HMI tags "DB_SDC_ERROR_STAT"
   "SDC\DB_SDC_ERROR_STAT\_Byte_DB_SDC_ERROR_STAT.F_STAT[XX5].EMS_TS_STAT_VAL.ERROR" : Int, internal   // Fehlernummer / Error number
   "SDC\DB_SDC_ERROR_STAT\_Byte_DB_SDC_ERROR_STAT.F_STAT[XX8].F" : Int, internal   // Fehler SDC + EMS Zusammenfassung / Fault SDC + EMS Summary
   "SDC\DB_SDC_ERROR_STAT\_Byte_DB_SDC_ERROR_STAT.F_STAT[X10].EMS_TS_STAT_VAL.DRIVE_POS_PERC" : Int, internal   // Position [% of Start End Section]
   "SDC\DB_SDC_ERROR_STAT\_Byte_DB_SDC_ERROR_STAT.F_STAT[XX9].F" : Int, internal   // Fehler SDC + EMS Zusammenfassung / Fault SDC + EMS Summary
   "SDC\DB_SDC_ERROR_STAT\_Byte_DB_SDC_ERROR_STAT.F_STAT[XX6].F_DATE" : Int, internal   // Fehler Zeit / Fault Time
   "SDC\DB_SDC_ERROR_STAT\DB_SDC_ERROR_STAT.F_STAT[XX7].EMS_TS_STAT_VAL.DRIVE_POS" : DInt AT %DB0.DBD0, 1 s   // Antriebsposition in mm / Drive position in mm
   "DB_SDC_ERRORS_STAT_HEADER.FAULT_PRO_SEITE_HMI" : Int = PLC DB_SDC_ERRORS_STAT.HEADER.FAULT_PRO_SEITE_HMI AT %DB3724.DBW10, 1 s   // Reserve
   "SDC\DB_SDC_ERROR_STAT\DB_SDC_ERROR_STAT.F_STAT[XX8].EMS_TS_STAT_VAL.DRIVE_POS" : DInt AT %DB0.DBD0, 1 s   // Antriebsposition in mm / Drive position in mm
   "SDC\DB_SDC_ERROR_STAT\DB_SDC_ERROR_STAT.F_STAT[XX8].EMS_TS_STAT_VAL.SEK" : Int AT %DB0.DBW0, 1 s   // Sektion
   "SDC\DB_SDC_ERROR_STAT\_Byte_DB_SDC_ERROR_STAT.F_STAT[XX1].EMS_TS_STAT_VAL.EMS_ID" : Int, internal   // EMS ID Nummer / EMS ID Number
   "SDC\DB_SDC_ERROR_STAT\DB_SDC_ERROR_STAT.F_STAT[XX5].EMS_TS_STAT_VAL.DRIVE_POS" : DInt AT %DB0.DBD0, 1 s   // Antriebsposition in mm / Drive position in mm
   "SDC\DB_SDC_ERROR_STAT\DB_SDC_ERROR_STAT.F_STAT[XX3].F_DATE" : Date_And_Time AT %DB0.DBX0.0, 1 s   // Fehler Zeit / Fault Time
   "SDC\DB_SDC_ERROR_STAT\_Byte_DB_SDC_ERROR_STAT.F_STAT[XX9].EMS_TS_STAT_VAL.TILT_POS" : Int, internal   // Tilt angle in degrees
   "SDC\DB_SDC_ERROR_STAT\DB_SDC_ERROR_STAT.F_STAT[XX7].F_DATE" : Date_And_Time AT %DB0.DBX0.0, 1 s   // Fehler Zeit / Fault Time
   "SDC\DB_SDC_ERROR_STAT\DB_SDC_ERROR_STAT.F_STAT[XX1].F_DATE" : Date_And_Time AT %DB0.DBX0.0, 1 s   // Fehler Zeit / Fault Time
   "SDC\DB_SDC_ERROR_STAT\DB_SDC_ERROR_STAT.F_STAT[XX4].EMS_TS_STAT_VAL.DRIVE_POS_PERC" : Int AT %DB0.DBW0, 1 s   // Position [% of Start End Section]
   "SDC\DB_SDC_ERROR_STAT\_Byte_DB_SDC_ERROR_STAT.F_STAT[XX6].EMS_TS_STAT_VAL.SEK" : Int, internal   // Sektion
   "SDC\DB_SDC_ERROR_STAT\_Byte_DB_SDC_ERROR_STAT.F_STAT[XX5].EMS_TS_STAT_VAL.PROFIL" : Int, internal   // Profile
   "SDC\DB_SDC_ERROR_STAT\DB_SDC_ERROR_STAT.F_STAT[XX5].EMS_TS_STAT_VAL.SEK" : Int AT %DB0.DBW0, 1 s   // Sektion
   "SDC\DB_SDC_ERROR_STAT\DB_SDC_ERROR_STAT.F_STAT[XX6].EMS_TS_STAT_VAL.PROFIL" : Int AT %DB0.DBW0, 1 s   // Profile
   "SDC\DB_SDC_ERROR_STAT\_Byte_DB_SDC_ERROR_STAT.F_STAT[XX8].EMS_TS_STAT_VAL.EMS_ID" : Int, internal   // EMS ID Nummer / EMS ID Number
   "SDC\DB_SDC_ERROR_STAT\_Byte_DB_SDC_ERROR_STAT.F_STAT[XX6].F" : Int, internal   // Fehler SDC + EMS Zusammenfassung / Fault SDC + EMS Summary
   "SDC\DB_SDC_ERROR_STAT\_Byte_DB_SDC_ERROR_STAT.F_STAT[XX5].EMS_TS_STAT_VAL.TILT_POS" : Int, internal   // Tilt angle in degrees
   "SDC\DB_SDC_ERROR_STAT\_Byte_DB_SDC_ERROR_STAT.F_STAT[XX2].EMS_TS_STAT_VAL.SEK" : Int, internal   // Sektion
   "SDC\DB_SDC_ERROR_STAT\DB_SDC_ERROR_STAT.F_STAT[XX5].F" : Word AT %DB0.DBW0, 1 s   // Fehler SDC + EMS Zusammenfassung / Fault SDC + EMS Summary
   "SDC\DB_SDC_ERROR_STAT\_Byte_DB_SDC_ERROR_STAT.F_STAT[XX7].F_DATE" : Int, internal   // Fehler Zeit / Fault Time
   "SDC\DB_SDC_ERROR_STAT\_Byte_DB_SDC_ERROR_STAT.F_STAT[XX6].EMS_TS_STAT_VAL.HOIST_POS" : Int, internal   // Höhe in mm / Height in mm
   "SDC\DB_SDC_ERROR_STAT\DB_SDC_ERROR_STAT.F_STAT[XX9].EMS_TS_STAT_VAL.HOIST_POS" : Int AT %DB0.DBW0, 1 s   // Höhe in mm / Height in mm
   "SDC\DB_SDC_ERROR_STAT\_Byte_DB_SDC_ERROR_STAT.F_STAT[XX1].EMS_TS_STAT_VAL.HOIST_POS" : Int, internal   // Höhe in mm / Height in mm
   "SDC\DB_SDC_ERROR_STAT\_Byte_DB_SDC_ERROR_STAT.F_STAT[XX5].EMS_TS_STAT_VAL.DRIVE_POS_PERC" : Int, internal   // Position [% of Start End Section]
   "SDC\DB_SDC_ERROR_STAT\DB_SDC_ERROR_STAT.F_STAT[XX1].EMS_TS_STAT_VAL.ERROR" : Int AT %DB0.DBW0, 1 s   // Fehlernummer / Error number
   "SDC\DB_SDC_ERROR_STAT\DB_SDC_ERROR_STAT.F_STAT[XX9].EMS_TS_STAT_VAL.SEK" : Int AT %DB0.DBW0, 1 s   // Sektion
   "SDC\DB_SDC_ERROR_STAT\_Byte_DB_SDC_ERROR_STAT.F_STAT[XX4].EMS_TS_STAT_VAL.DRIVE_POS" : Int, internal   // Antriebsposition in mm / Drive position in mm
   "SDC\DB_SDC_ERROR_STAT\DB_SDC_ERROR_STAT.F_STAT[XX4].EMS_TS_STAT_VAL.SEK" : Int AT %DB0.DBW0, 1 s   // Sektion
   "SDC\DB_SDC_ERROR_STAT\_Byte_DB_SDC_ERROR_STAT.F_STAT[XX2].F_DATE" : Int, internal   // Fehler Zeit / Fault Time
   "SDC\DB_SDC_ERROR_STAT\DB_SDC_ERROR_STAT.F_STAT[X10].EMS_TS_STAT_VAL.DRIVE_POS" : DInt AT %DB0.DBD0, 1 s   // Antriebsposition in mm / Drive position in mm
   "SDC\DB_SDC_ERROR_STAT\DB_SDC_ERROR_STAT.F_STAT[XX2].EMS_TS_STAT_VAL.TILT_POS" : Int AT %DB0.DBW0, 1 s   // Tilt angle in degrees
   "SDC\DB_SDC_ERROR_STAT\_Byte_DB_SDC_ERROR_STAT.F_STAT[XX2].EMS_TS_STAT_VAL.DRIVE_POS_PERC" : Int, internal   // Position [% of Start End Section]
   "SDC\DB_SDC_ERROR_STAT\_Byte_DB_SDC_ERROR_STAT.F_STAT[XX6].EMS_TS_STAT_VAL.TILT_POS" : Int, internal   // Tilt angle in degrees
   "SDC\DB_SDC_ERROR_STAT\DB_SDC_ERROR_STAT.F_STAT[XX5].EMS_TS_STAT_VAL.PROFIL" : Int AT %DB0.DBW0, 1 s   // Profile
   "SDC\DB_SDC_ERROR_STAT\_Byte_DB_SDC_ERROR_STAT.F_STAT[XX3].EMS_TS_STAT_VAL.EMS_ID" : Int, internal   // EMS ID Nummer / EMS ID Number
   "SDC\DB_SDC_ERROR_STAT\DB_SDC_ERROR_STAT.F_STAT[XX7].EMS_TS_STAT_VAL.SEK" : Int AT %DB0.DBW0, 1 s   // Sektion
   "SDC\DB_SDC_ERROR_STAT\DB_SDC_ERROR_STAT.F_STAT[XX1].EMS_TS_STAT_VAL.EMS_ID" : Int AT %DB0.DBW0, 1 s   // EMS ID Nummer / EMS ID Number
   "SDC\DB_SDC_ERROR_STAT\DB_SDC_ERROR_STAT.F_STAT[XX9].EMS_TS_STAT_VAL.TILT_POS" : Int AT %DB0.DBW0, 1 s   // Tilt angle in degrees
   "SDC\DB_SDC_ERROR_STAT\DB_SDC_ERROR_STAT.F_STAT[XX6].EMS_TS_STAT_VAL.HOIST_POS" : Int AT %DB0.DBW0, 1 s   // Höhe in mm / Height in mm
   "SDC\DB_SDC_ERROR_STAT\DB_SDC_ERROR_STAT.F_STAT[XX7].EMS_TS_STAT_VAL.PROFIL" : Int AT %DB0.DBW0, 1 s   // Profile
   "SDC\DB_SDC_ERROR_STAT\_Byte_DB_SDC_ERROR_STAT.F_STAT[XX8].EMS_TS_STAT_VAL.ERROR" : Int, internal   // Fehlernummer / Error number
   "SDC\DB_SDC_ERROR_STAT\DB_SDC_ERROR_STAT.F_STAT[XX3].EMS_TS_STAT_VAL.DRIVE_POS" : DInt AT %DB0.DBD0, 1 s   // Antriebsposition in mm / Drive position in mm
   "SDC\DB_SDC_ERROR_STAT\_Byte_DB_SDC_ERROR_STAT.F_STAT[XX9].EMS_TS_STAT_VAL.DRIVE_POS_PERC" : Int, internal   // Position [% of Start End Section]
   "SDC\DB_SDC_ERROR_STAT\_Byte_DB_SDC_ERROR_STAT.F_STAT[XX8].EMS_TS_STAT_VAL.DRIVE_POS_PERC" : Int, internal   // Position [% of Start End Section]
   "SDC\DB_SDC_ERROR_STAT\_Byte_DB_SDC_ERROR_STAT.F_STAT[X10].F" : Int, internal   // Fehler SDC + EMS Zusammenfassung / Fault SDC + EMS Summary
   "SDC\DB_SDC_ERROR_STAT\_Byte_DB_SDC_ERROR_STAT.F_STAT[XX9].EMS_TS_STAT_VAL.PROFIL" : Int, internal   // Profile
   "SDC\DB_SDC_ERROR_STAT\DB_SDC_ERROR_STAT.F_STAT[X10].EMS_TS_STAT_VAL.HOIST_POS" : Int AT %DB0.DBW0, 1 s   // Höhe in mm / Height in mm
   "SDC\DB_SDC_ERROR_STAT\DB_SDC_ERROR_STAT.F_STAT[X10].EMS_TS_STAT_VAL.SEK" : Int AT %DB0.DBW0, 1 s   // Sektion
   "SDC\DB_SDC_ERROR_STAT\_Byte_DB_SDC_ERROR_STAT.F_STAT[XX7].EMS_TS_STAT_VAL.SEK" : Int, internal   // Sektion
   "SDC\DB_SDC_ERROR_STAT\DB_SDC_ERROR_STAT.F_STAT[XX3].EMS_TS_STAT_VAL.PROFIL" : Int AT %DB0.DBW0, 1 s   // Profile
   "SDC\DB_SDC_ERROR_STAT\_Byte_DB_SDC_ERROR_STAT.F_STAT[XX4].F" : Int, internal   // Fehler SDC + EMS Zusammenfassung / Fault SDC + EMS Summary
   "SDC\DB_SDC_ERROR_STAT\_Byte_DB_SDC_ERROR_STAT.F_STAT[XX7].EMS_TS_STAT_VAL.ERROR" : Int, internal   // Fehlernummer / Error number
   "SDC\DB_SDC_ERROR_STAT\_intern_DB_Fault_Stat_Nr" : Int, internal
   "SDC\DB_SDC_ERROR_STAT\_Byte_DB_SDC_ERROR_STAT.F_STAT[XX6].EMS_TS_STAT_VAL.EMS_ID" : Int, internal   // EMS ID Nummer / EMS ID Number
   "SDC\DB_SDC_ERROR_STAT\_Byte_DB_SDC_ERROR_STAT.F_STAT[XX3].EMS_TS_STAT_VAL.DRIVE_POS_PERC" : Int, internal   // Position [% of Start End Section]
   "SDC\DB_SDC_ERROR_STAT\_Byte_DB_SDC_ERROR_STAT.F_STAT[XX6].EMS_TS_STAT_VAL.DRIVE_POS_PERC" : Int, internal   // Position [% of Start End Section]
   "SDC\DB_SDC_ERROR_STAT\_Byte_DB_SDC_ERROR_STAT.F_STAT[XX7].F" : Int, internal   // Fehler SDC + EMS Zusammenfassung / Fault SDC + EMS Summary
   "SDC\DB_SDC_ERROR_STAT\_Byte_DB_SDC_ERROR_STAT.F_STAT[X10].EMS_TS_STAT_VAL.ERROR" : Int, internal   // Fehlernummer / Error number
   "SDC\DB_SDC_ERROR_STAT\_Byte_DB_SDC_ERROR_STAT.F_STAT[XX2].EMS_TS_STAT_VAL.DRIVE_POS" : Int, internal   // Antriebsposition in mm / Drive position in mm
   "SDC\DB_SDC_ERROR_STAT\DB_SDC_ERROR_STAT.F_STAT[XX8].EMS_TS_STAT_VAL.ERROR" : Int AT %DB0.DBW0, 1 s   // Fehlernummer / Error number
   "SDC\DB_SDC_ERROR_STAT\DB_SDC_ERROR_STAT.F_STAT[XX7].EMS_TS_STAT_VAL.TILT_POS" : Int AT %DB0.DBW0, 1 s   // Tilt angle in degrees
   "DB_SDC_ERRORS_STAT_HEADER.MIN_NR_FAULT_STAT" : Int = PLC DB_SDC_ERRORS_STAT.HEADER.MIN_NR_FAULT_STAT AT %DB3724.DBW2, 1 s   // Niedrigste Fehler Nummer im Daten DB
   "SDC\DB_SDC_ERROR_STAT\DB_SDC_ERROR_STAT.F_STAT[XX2].EMS_TS_STAT_VAL.HOIST_POS" : Int AT %DB0.DBW0, 1 s   // Höhe in mm / Height in mm
   "SDC\DB_SDC_ERROR_STAT\DB_SDC_ERROR_STAT.F_STAT[XX5].EMS_TS_STAT_VAL.TILT_POS" : Int AT %DB0.DBW0, 1 s   // Tilt angle in degrees
   "SDC\DB_SDC_ERROR_STAT\DB_SDC_ERROR_STAT.F_STAT[XX2].F_DATE" : Date_And_Time AT %DB0.DBX0.0, 1 s   // Fehler Zeit / Fault Time
   "SDC\DB_SDC_ERROR_STAT\DB_SDC_ERROR_STAT.F_STAT[XX4].EMS_TS_STAT_VAL.HOIST_POS" : Int AT %DB0.DBW0, 1 s   // Höhe in mm / Height in mm
   "SDC\DB_SDC_ERROR_STAT\_Byte_DB_SDC_ERROR_STAT.F_STAT[XX5].EMS_TS_STAT_VAL.EMS_ID" : Int, internal   // EMS ID Nummer / EMS ID Number
   "SDC\DB_SDC_ERROR_STAT\DB_SDC_ERROR_STAT.F_STAT[XX8].F" : Word AT %DB0.DBW0, 1 s   // Fehler SDC + EMS Zusammenfassung / Fault SDC + EMS Summary
   "SDC\DB_SDC_ERROR_STAT\_Byte_DB_SDC_ERROR_STAT.F_STAT[XX7].EMS_TS_STAT_VAL.EMS_ID" : Int, internal   // EMS ID Nummer / EMS ID Number
   "SDC\DB_SDC_ERROR_STAT\DB_SDC_ERROR_STAT.F_STAT[XX2].EMS_TS_STAT_VAL.PROFIL" : Int AT %DB0.DBW0, 1 s   // Profile
   "SDC\DB_SDC_ERROR_STAT\DB_SDC_ERROR_STAT.F_STAT[XX1].EMS_TS_STAT_VAL.PROFIL" : Int AT %DB0.DBW0, 1 s   // Profile
   "SDC\DB_SDC_ERROR_STAT\_Byte_DB_SDC_ERROR_STAT.F_STAT[XX2].EMS_TS_STAT_VAL.PROFIL" : Int, internal   // Profile
   "SDC\DB_SDC_ERROR_STAT\_Byte_DB_SDC_ERROR_STAT.F_STAT[XX3].EMS_TS_STAT_VAL.ERROR" : Int, internal   // Fehlernummer / Error number
   "SDC\DB_SDC_ERROR_STAT\DB_SDC_ERROR_STAT.F_STAT[XX5].EMS_TS_STAT_VAL.ERROR" : Int AT %DB0.DBW0, 1 s   // Fehlernummer / Error number
   "SDC\DB_SDC_ERROR_STAT\_Byte_DB_SDC_ERROR_STAT.F_STAT[XX3].EMS_TS_STAT_VAL.TILT_POS" : Int, internal   // Tilt angle in degrees
   "SDC\DB_SDC_ERROR_STAT\_Byte_DB_SDC_ERROR_STAT.F_STAT[XX2].EMS_TS_STAT_VAL.ERROR" : Int, internal   // Fehlernummer / Error number
   "SDC\DB_SDC_ERROR_STAT\DB_SDC_ERROR_STAT.F_STAT[XX8].EMS_TS_STAT_VAL.HOIST_POS" : Int AT %DB0.DBW0, 1 s   // Höhe in mm / Height in mm
   "SDC\DB_SDC_ERROR_STAT\DB_SDC_ERROR_STAT.F_STAT[XX1].EMS_TS_STAT_VAL.DRIVE_POS_PERC" : Int AT %DB0.DBW0, 1 s   // Position [% of Start End Section]
   "SDC\DB_SDC_ERROR_STAT\DB_SDC_ERROR_STAT.F_STAT[XX9].EMS_TS_STAT_VAL.ERROR" : Int AT %DB0.DBW0, 1 s   // Fehlernummer / Error number
   "SDC\DB_SDC_ERROR_STAT\DB_SDC_ERROR_STAT.F_STAT[XX1].EMS_TS_STAT_VAL.TILT_POS" : Int AT %DB0.DBW0, 1 s   // Tilt angle in degrees
   "SDC\DB_SDC_ERROR_STAT\_Byte_DB_SDC_ERROR_STAT.F_STAT[XX1].EMS_TS_STAT_VAL.PROFIL" : Int, internal   // Profile
   "SDC\DB_SDC_ERROR_STAT\_Byte_DB_SDC_ERROR_STAT.F_STAT[XX4].EMS_TS_STAT_VAL.PROFIL" : Int, internal   // Profile
   "SDC\DB_SDC_ERROR_STAT\_Byte_DB_SDC_ERROR_STAT.F_STAT[XX1].EMS_TS_STAT_VAL.DRIVE_POS" : Int, internal   // Antriebsposition in mm / Drive position in mm
   "SDC\DB_SDC_ERROR_STAT\_Byte_DB_SDC_ERROR_STAT.F_STAT[XX7].EMS_TS_STAT_VAL.HOIST_POS" : Int, internal   // Höhe in mm / Height in mm
   "SDC\DB_SDC_ERROR_STAT\DB_SDC_ERROR_STAT.F_STAT[XX2].EMS_TS_STAT_VAL.DRIVE_POS_PERC" : Int AT %DB0.DBW0, 1 s   // Position [% of Start End Section]
   "SDC\DB_SDC_ERROR_STAT\_Byte_DB_SDC_ERROR_STAT.F_STAT[XX6].EMS_TS_STAT_VAL.PROFIL" : Int, internal   // Profile
   "DB_SDC_ERRORS_STAT_HEADER.START_FAULT_STAT" : Int = PLC DB_SDC_ERRORS_STAT.HEADER.START_FAULT_STAT AT %DB3724.DBW6, 1 s   // Startadresse der Fehler Daten im Daten DB
   "SDC\DB_SDC_ERROR_STAT\_Byte_DB_SDC_ERROR_STAT.F_STAT[X10].EMS_TS_STAT_VAL.EMS_ID" : Int, internal   // EMS ID Nummer / EMS ID Number
   "SDC\DB_SDC_ERROR_STAT\DB_SDC_ERROR_STAT.F_STAT[XX4].EMS_TS_STAT_VAL.ERROR" : Int AT %DB0.DBW0, 1 s   // Fehlernummer / Error number
   "SDC\DB_SDC_ERROR_STAT\DB_SDC_ERROR_STAT.F_STAT[XX6].EMS_TS_STAT_VAL.EMS_ID" : Int AT %DB0.DBW0, 1 s   // EMS ID Nummer / EMS ID Number
   "SDC\DB_SDC_ERROR_STAT\DB_SDC_ERROR_STAT.F_STAT[XX9].EMS_TS_STAT_VAL.DRIVE_POS_PERC" : Int AT %DB0.DBW0, 1 s   // Position [% of Start End Section]
   "SDC\DB_SDC_ERROR_STAT\_Byte_DB_SDC_ERROR_STAT.F_STAT[XX9].EMS_TS_STAT_VAL.HOIST_POS" : Int, internal   // Höhe in mm / Height in mm
   "SDC\DB_SDC_ERROR_STAT\DB_SDC_ERROR_STAT.F_STAT[XX9].F" : Word AT %DB0.DBW0, 1 s   // Fehler SDC + EMS Zusammenfassung / Fault SDC + EMS Summary
   "SDC\DB_SDC_ERROR_STAT\_Byte_DB_SDC_ERROR_STAT.F_STAT[XX1].F_DATE" : Int, internal   // Fehler Zeit / Fault Time
   "SDC\DB_SDC_ERROR_STAT\_Byte_DB_SDC_ERROR_STAT.F_STAT[XX9].EMS_TS_STAT_VAL.DRIVE_POS" : Int, internal   // Antriebsposition in mm / Drive position in mm
   "SDC\DB_SDC_ERROR_STAT\DB_SDC_ERROR_STAT.F_STAT[XX6].EMS_TS_STAT_VAL.ERROR" : Int AT %DB0.DBW0, 1 s   // Fehlernummer / Error number
   "SDC\DB_SDC_ERROR_STAT\DB_SDC_ERROR_STAT.F_STAT[XX3].EMS_TS_STAT_VAL.EMS_ID" : Int AT %DB0.DBW0, 1 s   // EMS ID Nummer / EMS ID Number
   "SDC\DB_SDC_ERROR_STAT\DB_SDC_ERROR_STAT.F_STAT[XX4].EMS_TS_STAT_VAL.PROFIL" : Int AT %DB0.DBW0, 1 s   // Profile
   "SDC\DB_SDC_ERROR_STAT\_Byte_DB_SDC_ERROR_STAT.F_STAT[XX3].EMS_TS_STAT_VAL.HOIST_POS" : Int, internal   // Höhe in mm / Height in mm
   "SDC\DB_SDC_ERROR_STAT\_Byte_DB_SDC_ERROR_STAT.F_STAT[XX1].EMS_TS_STAT_VAL.SEK" : Int, internal   // Sektion
   "SDC\DB_SDC_ERROR_STAT\_Byte_DB_SDC_ERROR_STAT.F_STAT[XX2].EMS_TS_STAT_VAL.EMS_ID" : Int, internal   // EMS ID Nummer / EMS ID Number
   "SDC\DB_SDC_ERROR_STAT\DB_SDC_ERROR_STAT.F_STAT[XX8].EMS_TS_STAT_VAL.PROFIL" : Int AT %DB0.DBW0, 1 s   // Profile
   "SDC\DB_SDC_ERROR_STAT\DB_SDC_ERROR_STAT.F_STAT[XX2].EMS_TS_STAT_VAL.SEK" : Int AT %DB0.DBW0, 1 s   // Sektion
   "SDC\DB_SDC_ERROR_STAT\_Byte_DB_SDC_ERROR_STAT.F_STAT[XX8].F_DATE" : Int, internal   // Fehler Zeit / Fault Time
   "SDC\DB_SDC_ERROR_STAT\DB_SDC_ERROR_STAT.F_STAT[XX9].F_DATE" : Date_And_Time AT %DB0.DBX0.0, 1 s   // Fehler Zeit / Fault Time
   "SDC\DB_SDC_ERROR_STAT\DB_SDC_ERROR_STAT.F_STAT[XX5].EMS_TS_STAT_VAL.HOIST_POS" : Int AT %DB0.DBW0, 1 s   // Höhe in mm / Height in mm
   "SDC\DB_SDC_ERROR_STAT\DB_SDC_ERROR_STAT.F_STAT[XX3].EMS_TS_STAT_VAL.ERROR" : Int AT %DB0.DBW0, 1 s   // Fehlernummer / Error number
   "SDC\DB_SDC_ERROR_STAT\DB_SDC_ERROR_STAT.F_STAT[XX6].F" : Word AT %DB0.DBW0, 1 s   // Fehler SDC + EMS Zusammenfassung / Fault SDC + EMS Summary
   "SDC\DB_SDC_ERROR_STAT\DB_SDC_ERROR_STAT.F_STAT[X10].EMS_TS_STAT_VAL.PROFIL" : Int AT %DB0.DBW0, 1 s   // Profile
   "DB_SDC_ERRORS_STAT_HEADER.LAENGE_FAULT_STAT" : Int = PLC DB_SDC_ERRORS_STAT.HEADER.LAENGE_FAULT_STAT AT %DB3724.DBW8, 1 s   // Länge Fehler Daten
   "SDC\DB_SDC_ERROR_STAT\DB_SDC_ERROR_STAT.F_STAT[XX2].EMS_TS_STAT_VAL.ERROR" : Int AT %DB0.DBW0, 1 s   // Fehlernummer / Error number
   "SDC\DB_SDC_ERROR_STAT\_Byte_DB_SDC_ERROR_STAT.F_STAT[X10].EMS_TS_STAT_VAL.DRIVE_POS" : Int, internal   // Antriebsposition in mm / Drive position in mm
   "SDC\DB_SDC_ERROR_STAT\_Byte_DB_SDC_ERROR_STAT.F_STAT[XX1].F" : Int, internal   // Fehler SDC + EMS Zusammenfassung / Fault SDC + EMS Summary
   "SDC\DB_SDC_ERROR_STAT\DB_SDC_ERROR_STAT.F_STAT[XX7].EMS_TS_STAT_VAL.DRIVE_POS_PERC" : Int AT %DB0.DBW0, 1 s
   "SDC\DB_SDC_ERROR_STAT\_Byte_DB_SDC_ERROR_STAT.F_STAT[XX4].EMS_TS_STAT_VAL.TILT_POS" : Int, internal   // Tilt angle in degrees
   "SDC\DB_SDC_ERROR_STAT\_Byte_DB_SDC_ERROR_STAT.F_STAT[XX5].F_DATE" : Int, internal   // Fehler Zeit / Fault Time
   "SDC\DB_SDC_ERROR_STAT\DB_SDC_ERROR_STAT.F_STAT[XX5].F_DATE" : Date_And_Time AT %DB0.DBX0.0, 1 s   // Fehler Zeit / Fault Time
   "SDC\DB_SDC_ERROR_STAT\_Byte_DB_SDC_ERROR_STAT.F_STAT[X10].EMS_TS_STAT_VAL.SEK" : Int, internal   // Sektion
   "SDC\DB_SDC_ERROR_STAT\DB_SDC_ERROR_STAT.F_STAT[XX7].EMS_TS_STAT_VAL.ERROR" : Int AT %DB0.DBW0, 1 s   // Fehlernummer / Error number
   "SDC\DB_SDC_ERROR_STAT\DB_SDC_ERROR_STAT.F_STAT[XX9].EMS_TS_STAT_VAL.DRIVE_POS" : DInt AT %DB0.DBD0, 1 s   // Antriebsposition in mm / Drive position in mm
   "SDC\DB_SDC_ERROR_STAT\_Byte_DB_SDC_ERROR_STAT.F_STAT[XX4].F_DATE" : Int, internal   // Fehler Zeit / Fault Time
   "SDC\DB_SDC_ERROR_STAT\_Byte_DB_SDC_ERROR_STAT.F_STAT[XX4].EMS_TS_STAT_VAL.DRIVE_POS_PERC" : Int, internal   // Position [% of Start End Section]
   "SDC\DB_SDC_ERROR_STAT\_Byte_DB_SDC_ERROR_STAT.F_STAT[XX4].EMS_TS_STAT_VAL.HOIST_POS" : Int, internal   // Höhe in mm / Height in mm
   "DB_SDC_ERRORS_STAT_HEADER.MAX_NR_FAULT_STAT" : Int = PLC DB_SDC_ERRORS_STAT.HEADER.MAX_NR_FAULT_STAT AT %DB3724.DBW4, 1 s   // Höchste Fehler Nummer im Daten DB
   "SDC\DB_SDC_ERROR_STAT\_Byte_DB_SDC_ERROR_STAT.F_STAT[XX7].EMS_TS_STAT_VAL.DRIVE_POS" : Int, internal   // Antriebsposition in mm / Drive position in mm
   "SDC\DB_SDC_ERROR_STAT\_Byte_DB_SDC_ERROR_STAT.F_STAT[X10].EMS_TS_STAT_VAL.HOIST_POS" : Int, internal   // Höhe in mm / Height in mm
   "SDC\DB_SDC_ERROR_STAT\_Byte_DB_SDC_ERROR_STAT.F_STAT[XX1].EMS_TS_STAT_VAL.DRIVE_POS_PERC" : Int, internal   // Position [% of Start End Section]
   "SDC\DB_SDC_ERROR_STAT\_Byte_DB_SDC_ERROR_STAT.F_STAT[XX7].EMS_TS_STAT_VAL.DRIVE_POS_PERC" : Int, internal   // Position [% of Start End Section]
   "SDC\DB_SDC_ERROR_STAT\DB_SDC_ERROR_STAT.F_STAT[XX1].EMS_TS_STAT_VAL.DRIVE_POS" : DInt AT %DB0.DBD0, 1 s   // Antriebsposition in mm / Drive position in mm
   "SDC\DB_SDC_ERROR_STAT\DB_SDC_ERROR_STAT.F_STAT[XX5].EMS_TS_STAT_VAL.DRIVE_POS_PERC" : Int AT %DB0.DBW0, 1 s   // Position [% of Start End Section]
   "SDC\DB_SDC_ERROR_STAT\_Byte_DB_SDC_ERROR_STAT.F_STAT[XX2].F" : Int, internal   // Fehler SDC + EMS Zusammenfassung / Fault SDC + EMS Summary
   "SDC\DB_SDC_ERROR_STAT\_Byte_DB_SDC_ERROR_STAT.F_STAT[XX2].EMS_TS_STAT_VAL.HOIST_POS" : Int, internal   // Höhe in mm / Height in mm
   "SDC\DB_SDC_ERROR_STAT\_Byte_DB_SDC_ERROR_STAT.F_STAT[X10].EMS_TS_STAT_VAL.TILT_POS" : Int, internal   // Tilt angle in degrees
   "SDC\DB_SDC_ERROR_STAT\_Byte_DB_SDC_ERROR_STAT.F_STAT[XX5].EMS_TS_STAT_VAL.DRIVE_POS" : Int, internal   // Antriebsposition in mm / Drive position in mm
   "SDC\DB_SDC_ERROR_STAT\DB_SDC_ERROR_STAT.F_STAT[XX4].EMS_TS_STAT_VAL.TILT_POS" : Int AT %DB0.DBW0, 1 s   // Tilt angle in degrees
   "SDC\DB_SDC_ERROR_STAT\_Byte_DB_SDC_ERROR_STAT.F_STAT[XX9].EMS_TS_STAT_VAL.EMS_ID" : Int, internal   // EMS ID Nummer / EMS ID Number
   "SDC\DB_SDC_ERROR_STAT\_Byte_DB_SDC_ERROR_STAT.F_STAT[X10].EMS_TS_STAT_VAL.PROFIL" : Int, internal   // Profile
   "SDC\DB_SDC_ERROR_STAT\_Byte_DB_SDC_ERROR_STAT.F_STAT[XX9].EMS_TS_STAT_VAL.ERROR" : Int, internal   // Fehlernummer / Error number
   "SDC\DB_SDC_ERROR_STAT\DB_SDC_ERROR_STAT.F_STAT[XX6].EMS_TS_STAT_VAL.TILT_POS" : Int AT %DB0.DBW0, 1 s   // Tilt angle in degrees
   "SDC\DB_SDC_ERROR_STAT\_Byte_DB_SDC_ERROR_STAT.F_STAT[XX5].EMS_TS_STAT_VAL.HOIST_POS" : Int, internal   // Höhe in mm / Height in mm
   "SDC\DB_SDC_ERROR_STAT\DB_SDC_ERROR_STAT.F_STAT[XX6].EMS_TS_STAT_VAL.DRIVE_POS" : DInt AT %DB0.DBD0, 1 s   // Antriebsposition in mm / Drive position in mm
   "SDC\DB_SDC_ERROR_STAT\DB_SDC_ERROR_STAT.F_STAT[XX4].F" : Word AT %DB0.DBW0, 1 s   // Fehler SDC + EMS Zusammenfassung / Fault SDC + EMS Summary
   "SDC\DB_SDC_ERROR_STAT\DB_SDC_ERROR_STAT.F_STAT[XX5].EMS_TS_STAT_VAL.EMS_ID" : Int AT %DB0.DBW0, 1 s   // EMS ID Nummer / EMS ID Number
   "SDC\DB_SDC_ERROR_STAT\DB_SDC_ERROR_STAT.F_STAT[XX8].F_DATE" : Date_And_Time AT %DB0.DBX0.0, 1 s   // Fehler Zeit / Fault Time
   "SDC\DB_SDC_ERROR_STAT\DB_SDC_ERROR_STAT.F_STAT[X10].EMS_TS_STAT_VAL.ERROR" : Int AT %DB0.DBW0, 1 s   // Fehlernummer / Error number
   "SDC\DB_SDC_ERROR_STAT\_Byte_DB_SDC_ERROR_STAT.F_STAT[XX1].EMS_TS_STAT_VAL.TILT_POS" : Int, internal   // Tilt angle in degrees
   "SDC\DB_SDC_ERROR_STAT\_Byte_DB_SDC_ERROR_STAT.F_STAT[XX8].EMS_TS_STAT_VAL.SEK" : Int, internal   // Sektion
   "SDC\DB_SDC_ERROR_STAT\DB_SDC_ERROR_STAT.F_STAT[XX7].EMS_TS_STAT_VAL.HOIST_POS" : Int AT %DB0.DBW0, 1 s   // Höhe in mm / Height in mm
   "SDC\DB_SDC_ERROR_STAT\DB_SDC_ERROR_STAT.F_STAT[XX2].EMS_TS_STAT_VAL.EMS_ID" : Int AT %DB0.DBW0, 1 s   // EMS ID Nummer / EMS ID Number
   "SDC\DB_SDC_ERROR_STAT\_Byte_DB_SDC_ERROR_STAT.F_STAT[XX9].EMS_TS_STAT_VAL.SEK" : Int, internal   // Sektion
   "SDC\DB_SDC_ERROR_STAT\_Byte_DB_SDC_ERROR_STAT.F_STAT[XX7].EMS_TS_STAT_VAL.TILT_POS" : Int, internal   // Tilt angle in degrees
   "SDC\DB_SDC_ERROR_STAT\_Byte_DB_SDC_ERROR_STAT.F_STAT[XX3].EMS_TS_STAT_VAL.DRIVE_POS" : Int, internal   // Antriebsposition in mm / Drive position in mm
   "SDC\DB_SDC_ERROR_STAT\DB_SDC_ERROR_STAT.F_STAT[XX9].EMS_TS_STAT_VAL.EMS_ID" : Int AT %DB0.DBW0, 1 s   // EMS ID Nummer / EMS ID Number
   "SDC\DB_SDC_ERROR_STAT\_intern_Fault_Stat_Nr_Array" : Array [0..9] of Int, internal
   "SDC\DB_SDC_ERROR_STAT\DB_SDC_ERROR_STAT.F_STAT[XX4].F_DATE" : Date_And_Time AT %DB0.DBX0.0, 1 s   // Fehler Zeit / Fault Time
   "SDC\DB_SDC_ERROR_STAT\DB_SDC_ERROR_STAT.F_STAT[XX4].EMS_TS_STAT_VAL.DRIVE_POS" : DInt AT %DB0.DBD0, 1 s   // Antriebsposition in mm / Drive position in mm
   "SDC\DB_SDC_ERROR_STAT\DB_SDC_ERROR_STAT.F_STAT[XX6].F_DATE" : Date_And_Time AT %DB0.DBX0.0, 1 s   // Fehler Zeit / Fault Time
   "SDC\DB_SDC_ERROR_STAT\DB_SDC_ERROR_STAT.F_STAT[XX2].EMS_TS_STAT_VAL.DRIVE_POS" : DInt AT %DB0.DBD0, 1 s   // Antriebsposition in mm / Drive position in mm
   "SDC\DB_SDC_ERROR_STAT\DB_SDC_ERROR_STAT.F_STAT[XX7].F" : Word AT %DB0.DBW0, 1 s   // Fehler SDC + EMS Zusammenfassung / Fault SDC + EMS Summary
   "SDC\DB_SDC_ERROR_STAT\_Byte_DB_SDC_ERROR_STAT.F_STAT[XX6].EMS_TS_STAT_VAL.DRIVE_POS" : Int, internal   // Antriebsposition in mm / Drive position in mm
   "SDC\DB_SDC_ERROR_STAT\DB_SDC_ERROR_STAT.F_STAT[X10].F_DATE" : Date_And_Time AT %DB0.DBX0.0, 1 s   // Fehler Zeit / Fault Time
   "SDC\DB_SDC_ERROR_STAT\_Byte_DB_SDC_ERROR_STAT.F_STAT[XX9].F_DATE" : Int, internal   // Fehler Zeit / Fault Time
   "SDC\DB_SDC_ERROR_STAT\DB_SDC_ERROR_STAT.F_STAT[X10].EMS_TS_STAT_VAL.TILT_POS" : Int AT %DB0.DBW0, 1 s   // Tilt angle in degrees
   "SDC\DB_SDC_ERROR_STAT\_Byte_DB_SDC_ERROR_STAT.F_STAT[XX8].EMS_TS_STAT_VAL.TILT_POS" : Int, internal   // Tilt angle in degrees
   "SDC\DB_SDC_ERROR_STAT\DB_SDC_ERROR_STAT.F_STAT[XX2].F" : Word AT %DB0.DBW0, 1 s   // Fehler SDC + EMS Zusammenfassung / Fault SDC + EMS Summary
   "SDC\DB_SDC_ERROR_STAT\_Byte_DB_SDC_ERROR_STAT.F_STAT[XX3].F_DATE" : Int, internal   // Fehler Zeit / Fault Time
   "SDC\DB_SDC_ERROR_STAT\DB_SDC_ERROR_STAT.F_STAT[XX8].EMS_TS_STAT_VAL.TILT_POS" : Int AT %DB0.DBW0, 1 s   // Tilt angle in degrees
   "SDC\DB_SDC_ERROR_STAT\DB_SDC_ERROR_STAT.F_STAT[X10].EMS_TS_STAT_VAL.DRIVE_POS_PERC" : Int AT %DB0.DBW0, 1 s   // Position [% of Start End Section]
   "SDC\DB_SDC_ERROR_STAT\DB_SDC_ERROR_STAT.F_STAT[XX6].EMS_TS_STAT_VAL.DRIVE_POS_PERC" : Int AT %DB0.DBW0, 1 s   // Position [% of Start End Section]
   "SDC\DB_SDC_ERROR_STAT\DB_SDC_ERROR_STAT.F_STAT[X10].EMS_TS_STAT_VAL.EMS_ID" : Int AT %DB0.DBW0, 1 s   // EMS ID Nummer / EMS ID Number
   "SDC\DB_SDC_ERROR_STAT\_Byte_DB_SDC_ERROR_STAT.F_STAT[XX2].EMS_TS_STAT_VAL.TILT_POS" : Int, internal   // Tilt angle in degrees
   "SDC\DB_SDC_ERROR_STAT\DB_SDC_ERROR_STAT.F_STAT[XX7].EMS_TS_STAT_VAL.EMS_ID" : Int AT %DB0.DBW0, 1 s   // EMS ID Nummer / EMS ID Number
   "SDC\DB_SDC_ERROR_STAT\DB_SDC_ERROR_STAT.F_STAT[XX1].EMS_TS_STAT_VAL.SEK" : Int AT %DB0.DBW0, 1 s   // Sektion
   "SDC\DB_SDC_ERROR_STAT\_Byte_DB_SDC_ERROR_STAT.F_STAT[XX8].EMS_TS_STAT_VAL.DRIVE_POS" : Int, internal   // Antriebsposition in mm / Drive position in mm
   "SDC\DB_SDC_ERROR_STAT\_Byte_DB_SDC_ERROR_STAT.F_STAT[XX7].EMS_TS_STAT_VAL.PROFIL" : Int, internal   // Profile
   "SDC\DB_SDC_ERROR_STAT\_Byte_DB_SDC_ERROR_STAT.F_STAT[XX3].EMS_TS_STAT_VAL.SEK" : Int, internal   // Sektion
   "SDC\DB_SDC_ERROR_STAT\DB_SDC_ERROR_STAT.F_STAT[XX8].EMS_TS_STAT_VAL.EMS_ID" : Int AT %DB0.DBW0, 1 s   // EMS ID Nummer / EMS ID Number
   "SDC\DB_SDC_ERROR_STAT\DB_SDC_ERROR_STAT.F_STAT[XX4].EMS_TS_STAT_VAL.EMS_ID" : Int AT %DB0.DBW0, 1 s   // EMS ID Nummer / EMS ID Number
   "SDC\DB_SDC_ERROR_STAT\DB_SDC_ERROR_STAT.F_STAT[XX3].EMS_TS_STAT_VAL.SEK" : Int AT %DB0.DBW0, 1 s   // Sektion
   "DB_SDC_ERRORS_STAT_HEADER.DB_NR" : Int = PLC DB_SDC_ERRORS_STAT.HEADER.DB_NR AT %DB3724.DBW0, 1 s   // DB Nummer
   "SDC\DB_SDC_ERROR_STAT\_Byte_DB_SDC_ERROR_STAT.F_STAT[XX6].EMS_TS_STAT_VAL.ERROR" : Int, internal   // Fehlernummer / Error number
   "SDC\DB_SDC_ERROR_STAT\_Byte_DB_SDC_ERROR_STAT.F_STAT[XX8].EMS_TS_STAT_VAL.PROFIL" : Int, internal   // Profile
   "SDC\DB_SDC_ERROR_STAT\DB_SDC_ERROR_STAT.F_STAT[XX1].F" : Word AT %DB0.DBW0, 1 s   // Fehler SDC + EMS Zusammenfassung / Fault SDC + EMS Summary
   "SDC\DB_SDC_ERROR_STAT\DB_SDC_ERROR_STAT.F_STAT[XX1].EMS_TS_STAT_VAL.HOIST_POS" : Int AT %DB0.DBW0, 1 s   // Höhe in mm / Height in mm
   "SDC\DB_SDC_ERROR_STAT\_Byte_DB_SDC_ERROR_STAT.F_STAT[XX4].EMS_TS_STAT_VAL.ERROR" : Int, internal   // Fehlernummer / Error number
   "SDC\DB_SDC_ERROR_STAT\_Byte_DB_SDC_ERROR_STAT.F_STAT[X10].F_DATE" : Int, internal   // Fehler Zeit / Fault Time
   "SDC\DB_SDC_ERROR_STAT\_Byte_DB_SDC_ERROR_STAT.F_STAT[XX4].EMS_TS_STAT_VAL.EMS_ID" : Int, internal   // EMS ID Nummer / EMS ID Number
   "SDC\DB_SDC_ERROR_STAT\DB_SDC_ERROR_STAT.F_STAT[XX3].EMS_TS_STAT_VAL.TILT_POS" : Int AT %DB0.DBW0, 1 s   // Tilt angle in degrees
   "SDC\DB_SDC_ERROR_STAT\_Byte_DB_SDC_ERROR_STAT.F_STAT[XX4].EMS_TS_STAT_VAL.SEK" : Int, internal   // Sektion
   "SDC\DB_SDC_ERROR_STAT\_Byte_DB_SDC_ERROR_STAT.F_STAT[XX3].EMS_TS_STAT_VAL.PROFIL" : Int, internal   // Profile
   "SDC\DB_SDC_ERROR_STAT\_Byte_DB_SDC_ERROR_STAT.F_STAT[XX5].EMS_TS_STAT_VAL.SEK" : Int, internal   // Sektion
   "SDC\DB_SDC_ERROR_STAT\_Byte_DB_SDC_ERROR_STAT.F_STAT[XX8].EMS_TS_STAT_VAL.HOIST_POS" : Int, internal   // Höhe in mm / Height in mm
   "SDC\DB_SDC_ERROR_STAT\_intern_Fault_Stat_Nr" : Int, internal
   "SDC\DB_SDC_ERROR_STAT\DB_SDC_ERROR_STAT.F_STAT[X10].F" : Word AT %DB0.DBW0, 1 s   // Fehler SDC + EMS Zusammenfassung / Fault SDC + EMS Summary
   "SDC\DB_SDC_ERROR_STAT\DB_SDC_ERROR_STAT.F_STAT[XX8].EMS_TS_STAT_VAL.DRIVE_POS_PERC" : Int AT %DB0.DBW0, 1 s   // Position [% of Start End Section]
   "SDC\DB_SDC_ERROR_STAT\DB_SDC_ERROR_STAT.F_STAT[XX9].EMS_TS_STAT_VAL.PROFIL" : Int AT %DB0.DBW0, 1 s   // Profile
   "SDC\DB_SDC_ERROR_STAT\DB_SDC_ERROR_STAT.F_STAT[XX3].EMS_TS_STAT_VAL.HOIST_POS" : Int AT %DB0.DBW0, 1 s   // Höhe in mm / Height in mm
   "SDC\DB_SDC_ERROR_STAT\DB_SDC_ERROR_STAT.F_STAT[XX3].F" : Word AT %DB0.DBW0, 1 s   // Fehler SDC + EMS Zusammenfassung / Fault SDC + EMS Summary
   "SDC\DB_SDC_ERROR_STAT\DB_SDC_ERROR_STAT.F_STAT[XX3].EMS_TS_STAT_VAL.DRIVE_POS_PERC" : Int AT %DB0.DBW0, 1 s   // Position [% of Start End Section]
   "SDC\DB_SDC_ERROR_STAT\_Byte_DB_SDC_ERROR_STAT.F_STAT[XX3].F" : Int, internal   // Fehler SDC + EMS Zusammenfassung / Fault SDC + EMS Summary
   "SDC\DB_SDC_ERROR_STAT\_Byte_DB_SDC_ERROR_STAT.F_STAT[XX1].EMS_TS_STAT_VAL.ERROR" : Int, internal   // Fehlernummer / Error number
   "SDC\DB_SDC_ERROR_STAT\_Byte_DB_SDC_ERROR_STAT.F_STAT[XX5].F" : Int, internal   // Fehler SDC + EMS Zusammenfassung / Fault SDC + EMS Summary
   "SDC\DB_SDC_ERROR_STAT\DB_SDC_ERROR_STAT.F_STAT[XX6].EMS_TS_STAT_VAL.SEK" : Int AT %DB0.DBW0, 1 s   // Sektion
   "DB_SDC_ERRORS_STAT_HEADER.RESET_ARCH" : Bool = PLC DB_SDC_ERRORS_STAT.HEADER.RESET_ARCH AT %DB3724.DBX18.1, 1 s

HMI tags "DB_SDC_ERROR_STAT_EMS001"
   "DB_SDC_ERRORS_STAT_ER_AKT[1].ER_TRIGER" : Word = PLC DB_SDC_ERRORS_STAT.ER_AKT[1].ER_TRIGER AT %DB3724.DBW28020, 1 s
   "DB_SDC_ERRORS_STAT_ER_AKT[1].ER_STAT[1].DRIVE_POS" : DInt = PLC DB_SDC_ERRORS_STAT.ER_AKT[1].ER_STAT[1].DRIVE_POS AT %DB3724.DBD28026, 1 s
   "DB_SDC_ERRORS_STAT_ER_AKT[1].ER_STAT[1].ERROR" : Int = PLC DB_SDC_ERRORS_STAT.ER_AKT[1].ER_STAT[1].ERROR AT %DB3724.DBW28032, 1 s
   "DB_SDC_ERRORS_STAT_ER_AKT[1].ER_STAT[2].DRIVE_POS" : DInt = PLC DB_SDC_ERRORS_STAT.ER_AKT[1].ER_STAT[2].DRIVE_POS AT %DB3724.DBD28042, 1 s
   "DB_SDC_ERRORS_STAT_ER_AKT[1].ER_STAT[2].ERROR" : Int = PLC DB_SDC_ERRORS_STAT.ER_AKT[1].ER_STAT[2].ERROR AT %DB3724.DBW28048, 1 s
   "DB_SDC_ERRORS_STAT_ER_AKT[1].ER_STAT[3].DRIVE_POS" : DInt = PLC DB_SDC_ERRORS_STAT.ER_AKT[1].ER_STAT[3].DRIVE_POS AT %DB3724.DBD28058, 1 s
   "DB_SDC_ERRORS_STAT_ER_AKT[1].ER_STAT[3].ERROR" : Int = PLC DB_SDC_ERRORS_STAT.ER_AKT[1].ER_STAT[3].ERROR AT %DB3724.DBW28064, 1 s
   "DB_SDC_ERRORS_STAT_ER_AKT[1].ER_STAT[4].DRIVE_POS" : DInt = PLC DB_SDC_ERRORS_STAT.ER_AKT[1].ER_STAT[4].DRIVE_POS AT %DB3724.DBD28074, 1 s
   "DB_SDC_ERRORS_STAT_ER_AKT[1].ER_STAT[4].ERROR" : Int = PLC DB_SDC_ERRORS_STAT.ER_AKT[1].ER_STAT[4].ERROR AT %DB3724.DBW28080, 1 s

HMI tags "DB_SDC_ERROR_STAT_EMS002"
   "DB_SDC_ERRORS_STAT_ER_AKT[2].ER_TRIGER" : Word = PLC DB_SDC_ERRORS_STAT.ER_AKT[2].ER_TRIGER AT %DB3724.DBW28086, 1 s
   "DB_SDC_ERRORS_STAT_ER_AKT[2].ER_STAT[1].DRIVE_POS" : DInt = PLC DB_SDC_ERRORS_STAT.ER_AKT[2].ER_STAT[1].DRIVE_POS AT %DB3724.DBD28092, 1 s
   "DB_SDC_ERRORS_STAT_ER_AKT[2].ER_STAT[1].ERROR" : Int = PLC DB_SDC_ERRORS_STAT.ER_AKT[2].ER_STAT[1].ERROR AT %DB3724.DBW28098, 1 s
   "DB_SDC_ERRORS_STAT_ER_AKT[2].ER_STAT[2].DRIVE_POS" : DInt = PLC DB_SDC_ERRORS_STAT.ER_AKT[2].ER_STAT[2].DRIVE_POS AT %DB3724.DBD28108, 1 s
   "DB_SDC_ERRORS_STAT_ER_AKT[2].ER_STAT[2].ERROR" : Int = PLC DB_SDC_ERRORS_STAT.ER_AKT[2].ER_STAT[2].ERROR AT %DB3724.DBW28114, 1 s
   "DB_SDC_ERRORS_STAT_ER_AKT[2].ER_STAT[3].DRIVE_POS" : DInt = PLC DB_SDC_ERRORS_STAT.ER_AKT[2].ER_STAT[3].DRIVE_POS AT %DB3724.DBD28124, 1 s
   "DB_SDC_ERRORS_STAT_ER_AKT[2].ER_STAT[3].ERROR" : Int = PLC DB_SDC_ERRORS_STAT.ER_AKT[2].ER_STAT[3].ERROR AT %DB3724.DBW28130, 1 s
   "DB_SDC_ERRORS_STAT_ER_AKT[2].ER_STAT[4].DRIVE_POS" : DInt = PLC DB_SDC_ERRORS_STAT.ER_AKT[2].ER_STAT[4].DRIVE_POS AT %DB3724.DBD28140, 1 s
   "DB_SDC_ERRORS_STAT_ER_AKT[2].ER_STAT[4].ERROR" : Int = PLC DB_SDC_ERRORS_STAT.ER_AKT[2].ER_STAT[4].ERROR AT %DB3724.DBW28146, 1 s

HMI tags "DB_SDC_ERROR_STAT_EMS003"
   "DB_SDC_ERRORS_STAT_ER_AKT[3].ER_TRIGER" : Word = PLC DB_SDC_ERRORS_STAT.ER_AKT[3].ER_TRIGER AT %DB3724.DBW28152, 1 s
   "DB_SDC_ERRORS_STAT_ER_AKT[3].ER_STAT[1].DRIVE_POS" : DInt = PLC DB_SDC_ERRORS_STAT.ER_AKT[3].ER_STAT[1].DRIVE_POS AT %DB3724.DBD28158, 1 s
   "DB_SDC_ERRORS_STAT_ER_AKT[3].ER_STAT[1].ERROR" : Int = PLC DB_SDC_ERRORS_STAT.ER_AKT[3].ER_STAT[1].ERROR AT %DB3724.DBW28164, 1 s
   "DB_SDC_ERRORS_STAT_ER_AKT[3].ER_STAT[2].DRIVE_POS" : DInt = PLC DB_SDC_ERRORS_STAT.ER_AKT[3].ER_STAT[2].DRIVE_POS AT %DB3724.DBD28174, 1 s
   "DB_SDC_ERRORS_STAT_ER_AKT[3].ER_STAT[2].ERROR" : Int = PLC DB_SDC_ERRORS_STAT.ER_AKT[3].ER_STAT[2].ERROR AT %DB3724.DBW28180, 1 s
   "DB_SDC_ERRORS_STAT_ER_AKT[3].ER_STAT[3].DRIVE_POS" : DInt = PLC DB_SDC_ERRORS_STAT.ER_AKT[3].ER_STAT[3].DRIVE_POS AT %DB3724.DBD28190, 1 s
   "DB_SDC_ERRORS_STAT_ER_AKT[3].ER_STAT[3].ERROR" : Int = PLC DB_SDC_ERRORS_STAT.ER_AKT[3].ER_STAT[3].ERROR AT %DB3724.DBW28196, 1 s
   "DB_SDC_ERRORS_STAT_ER_AKT[3].ER_STAT[4].DRIVE_POS" : DInt = PLC DB_SDC_ERRORS_STAT.ER_AKT[3].ER_STAT[4].DRIVE_POS AT %DB3724.DBD28206, 1 s
   "DB_SDC_ERRORS_STAT_ER_AKT[3].ER_STAT[4].ERROR" : Int = PLC DB_SDC_ERRORS_STAT.ER_AKT[3].ER_STAT[4].ERROR AT %DB3724.DBW28212, 1 s

HMI tags "DB_SDC_ERROR_STAT_EMS004"
   "DB_SDC_ERRORS_STAT_ER_AKT[4].ER_TRIGER" : Word = PLC DB_SDC_ERRORS_STAT.ER_AKT[4].ER_TRIGER AT %DB3724.DBW28218, 1 s
   "DB_SDC_ERRORS_STAT_ER_AKT[4].ER_STAT[1].DRIVE_POS" : DInt = PLC DB_SDC_ERRORS_STAT.ER_AKT[4].ER_STAT[1].DRIVE_POS AT %DB3724.DBD28224, 1 s
   "DB_SDC_ERRORS_STAT_ER_AKT[4].ER_STAT[1].ERROR" : Int = PLC DB_SDC_ERRORS_STAT.ER_AKT[4].ER_STAT[1].ERROR AT %DB3724.DBW28230, 1 s
   "DB_SDC_ERRORS_STAT_ER_AKT[4].ER_STAT[2].DRIVE_POS" : DInt = PLC DB_SDC_ERRORS_STAT.ER_AKT[4].ER_STAT[2].DRIVE_POS AT %DB3724.DBD28240, 1 s
   "DB_SDC_ERRORS_STAT_ER_AKT[4].ER_STAT[2].ERROR" : Int = PLC DB_SDC_ERRORS_STAT.ER_AKT[4].ER_STAT[2].ERROR AT %DB3724.DBW28246, 1 s
   "DB_SDC_ERRORS_STAT_ER_AKT[4].ER_STAT[3].DRIVE_POS" : DInt = PLC DB_SDC_ERRORS_STAT.ER_AKT[4].ER_STAT[3].DRIVE_POS AT %DB3724.DBD28256, 1 s
   "DB_SDC_ERRORS_STAT_ER_AKT[4].ER_STAT[3].ERROR" : Int = PLC DB_SDC_ERRORS_STAT.ER_AKT[4].ER_STAT[3].ERROR AT %DB3724.DBW28262, 1 s
   "DB_SDC_ERRORS_STAT_ER_AKT[4].ER_STAT[4].DRIVE_POS" : DInt = PLC DB_SDC_ERRORS_STAT.ER_AKT[4].ER_STAT[4].DRIVE_POS AT %DB3724.DBD28272, 1 s
   "DB_SDC_ERRORS_STAT_ER_AKT[4].ER_STAT[4].ERROR" : Int = PLC DB_SDC_ERRORS_STAT.ER_AKT[4].ER_STAT[4].ERROR AT %DB3724.DBW28278, 1 s
